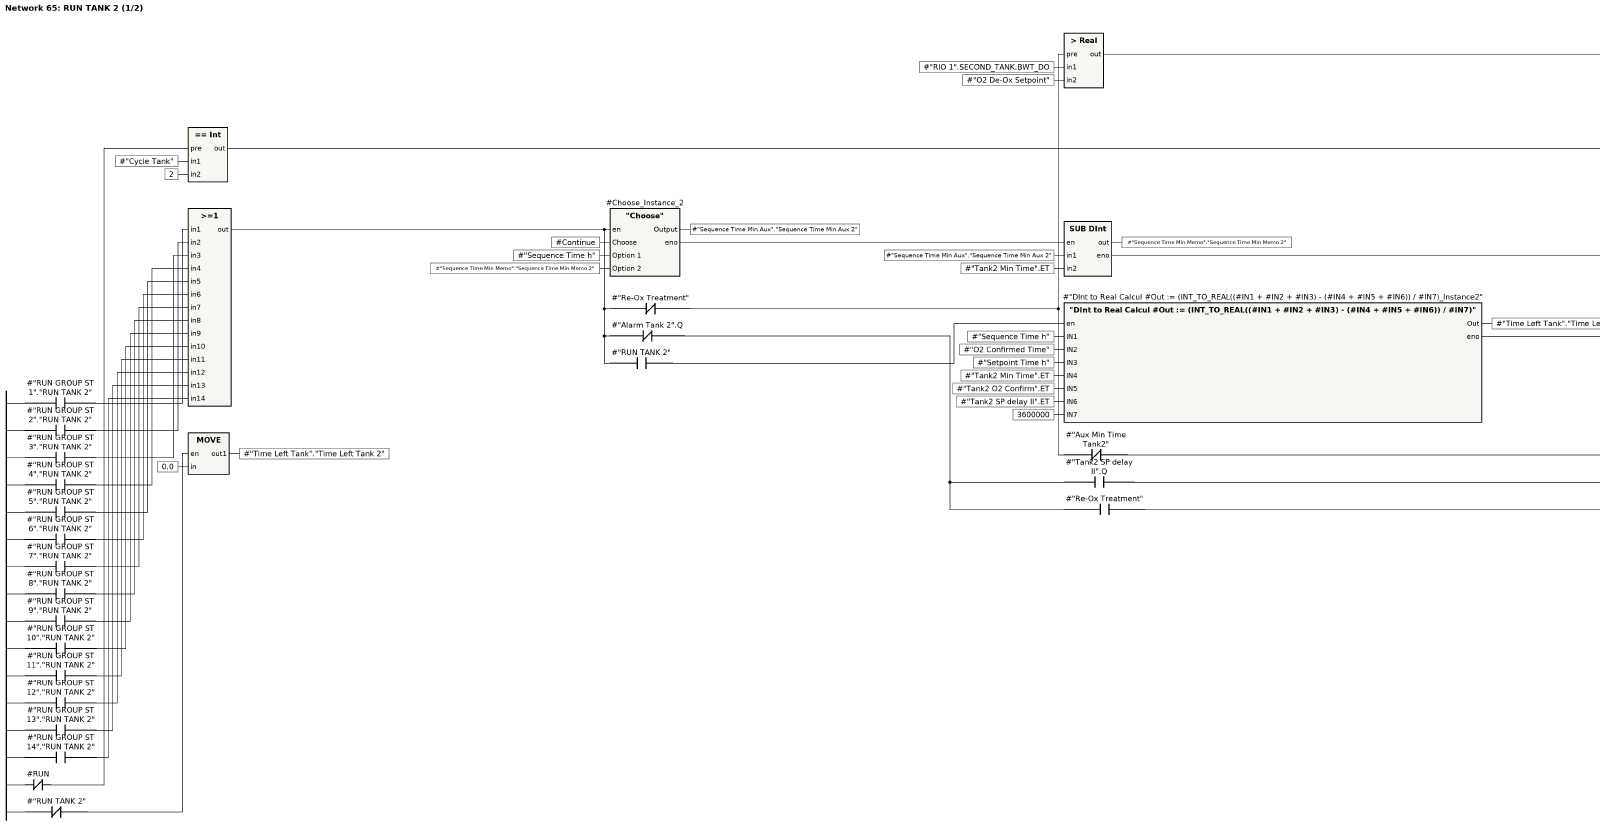
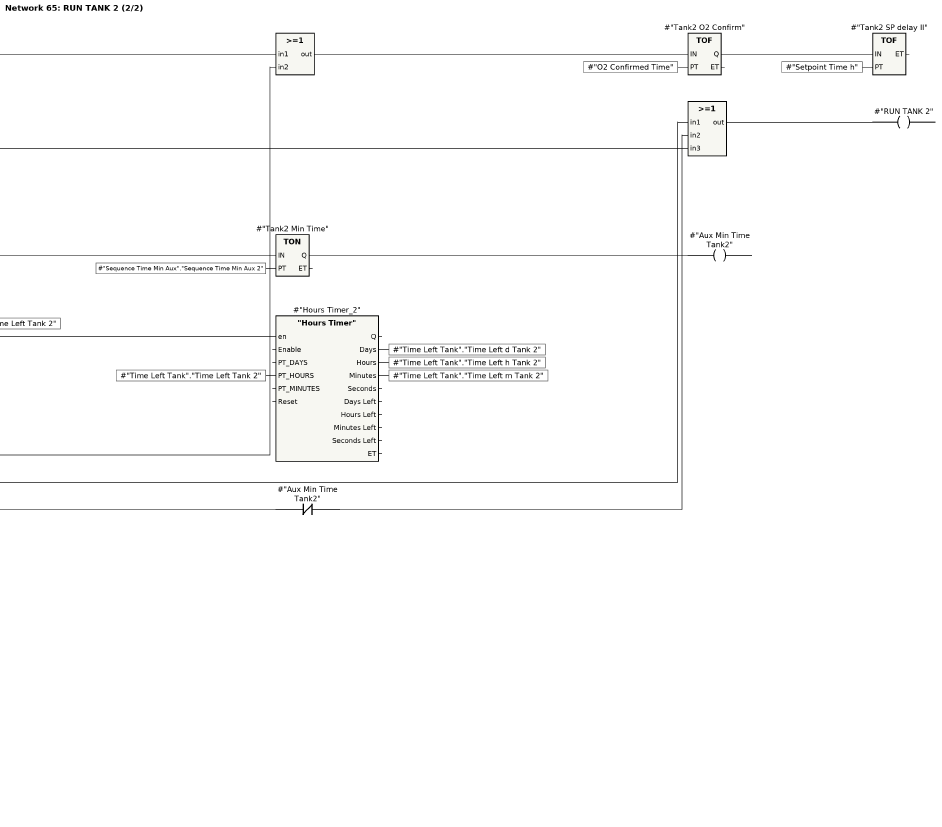
   #_w1 := #"RUN GROUP ST 1"."RUN TANK 2" OR #"RUN GROUP ST 2"."RUN TANK 2" OR #"RUN GROUP ST 3"."RUN TANK 2" OR #"RUN GROUP ST 4"."RUN TANK 2" OR #"RUN GROUP ST 5"."RUN TANK 2" OR #"RUN GROUP ST 6"."RUN TANK 2" OR #"RUN GROUP ST 7"."RUN TANK 2" OR #"RUN GROUP ST 8"."RUN TANK 2" OR #"RUN GROUP ST 9"."RUN TANK 2" OR #"RUN GROUP ST 10"."RUN TANK 2" OR #"RUN GROUP ST 11"."RUN TANK 2" OR #"RUN GROUP ST 12"."RUN TANK 2" OR #"RUN GROUP ST 13"."RUN TANK 2" OR #"RUN GROUP ST 14"."RUN TANK 2";
   #Choose_Instance_2(EN := #_w1,   // "Choose"
                      Choose := #Continue,
                      "Option 1" := #"Sequence Time h",
                      "Option 2" := #"Sequence Time Min Memo"."Sequence Time Min Memo 2",
                      Output => #"Sequence Time Min Aux"."Sequence Time Min Aux 2",
                      ENO => #_w2);
   IF #_w2 THEN
       #"Sequence Time Min Memo"."Sequence Time Min Memo 2" := #"Sequence Time Min Aux"."Sequence Time Min Aux 2" - #"Tank2 Min Time".ET;
   END_IF;
   #"Tank2 Min Time"(IN := #_w2, PT := #"Sequence Time Min Aux"."Sequence Time Min Aux 2");   // TON
   #"Aux Min Time Tank2" := #"Tank2 Min Time".Q;
   #"Tank2 O2 Confirm"(IN := #_w1 AND NOT #"Re-Ox Treatment" AND ((#"RIO 1".SECOND_TANK.BWT_DO > #"O2 De-Ox Setpoint") OR NOT #"Aux Min Time Tank2"),   // TOF
                       PT := #"O2 Confirmed Time");
   #"Tank2 SP delay II"(IN := #"Tank2 O2 Confirm".Q, PT := #"Setpoint Time h");   // TOF
   #"DInt to Real Calcul #Out := (INT_TO_REAL((#IN1 + #IN2 + #IN3) - (#IN4 + #IN5 + #IN6)) / #IN7)_Instance2"(EN := #_w1 AND #"RUN TANK 2",   // "DInt to Real Calcul #Out := (INT_TO_REAL((#IN1 + #IN2 + #IN3) - (#IN4 + #IN5 + #IN6)) / #IN7)"
                           IN1 := #"Sequence Time h",
                           IN2 := #"O2 Confirmed Time",
                           IN3 := #"Setpoint Time h",
                           IN4 := #"Tank2 Min Time".ET,
                           IN5 := #"Tank2 O2 Confirm".ET,
                           IN6 := #"Tank2 SP delay II".ET,
                           IN7 := 3600000,
                           Out => #"Time Left Tank"."Time Left Tank 2",
                           ENO => #_w3);
   IF #_w3 THEN
       #"Hours Timer_2"(PT_HOURS := #"Time Left Tank"."Time Left Tank 2",   // "Hours Timer"
                        Days => #"Time Left Tank"."Time Left d Tank 2",
                        Hours => #"Time Left Tank"."Time Left h Tank 2",
                        Minutes => #"Time Left Tank"."Time Left m Tank 2");
   END_IF;
   #"RUN TANK 2" := (#_w1 AND NOT #"Alarm Tank 2".Q AND (#"Tank2 SP delay II".Q OR (#"Re-Ox Treatment" AND NOT #"Aux Min Time Tank2"))) OR (NOT #RUN AND (#"Cycle Tank" = 2));
   IF NOT #"RUN TANK 2" THEN #"Time Left Tank"."Time Left Tank 2" := 0.0; END_IF;
END_REGION

REGION Network 66: RUN TANK 3
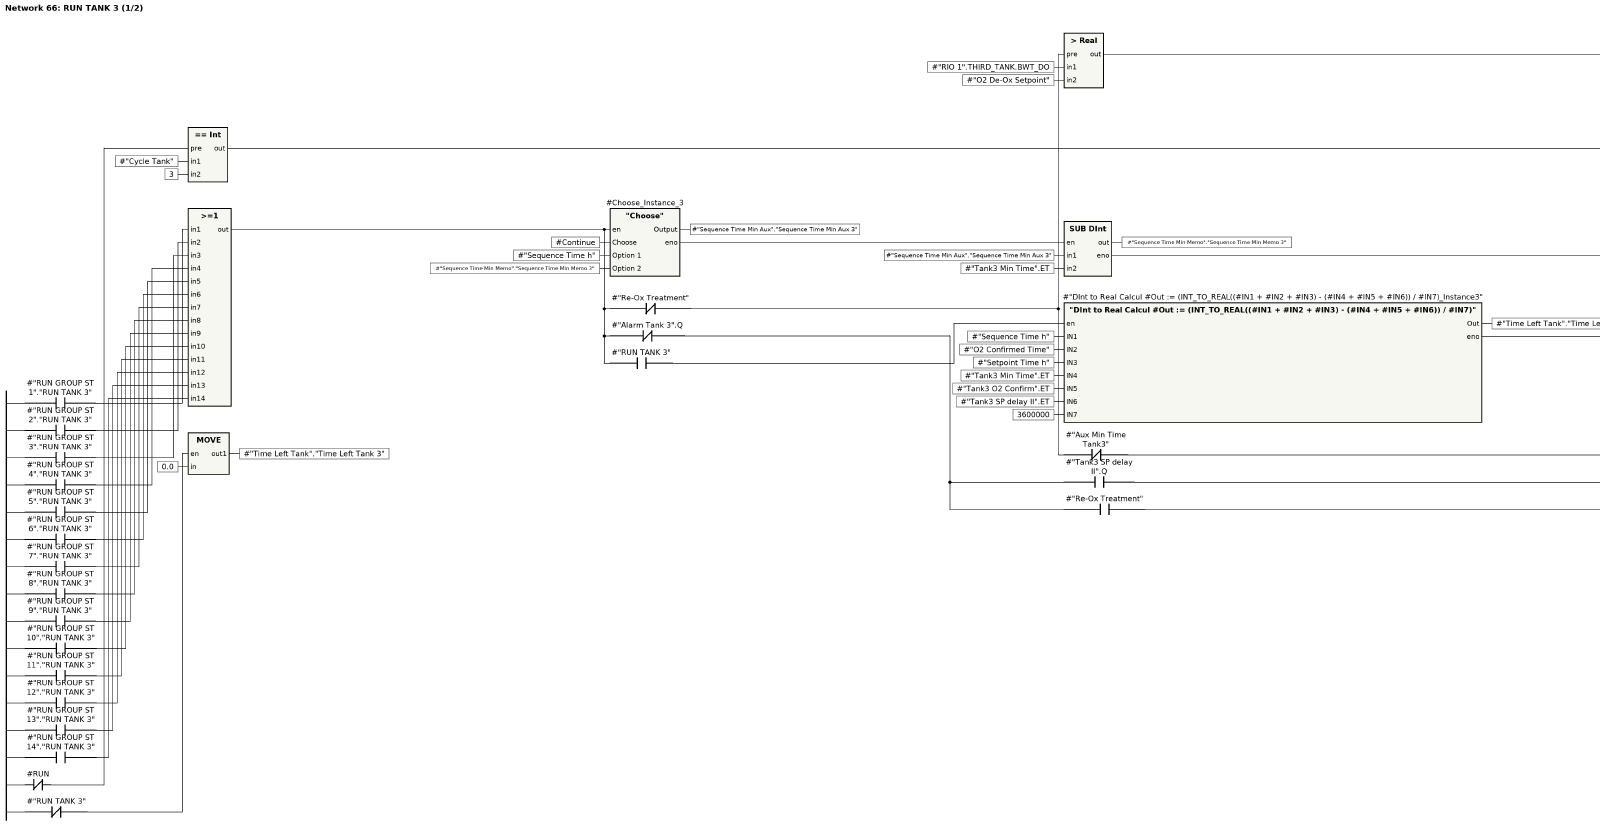
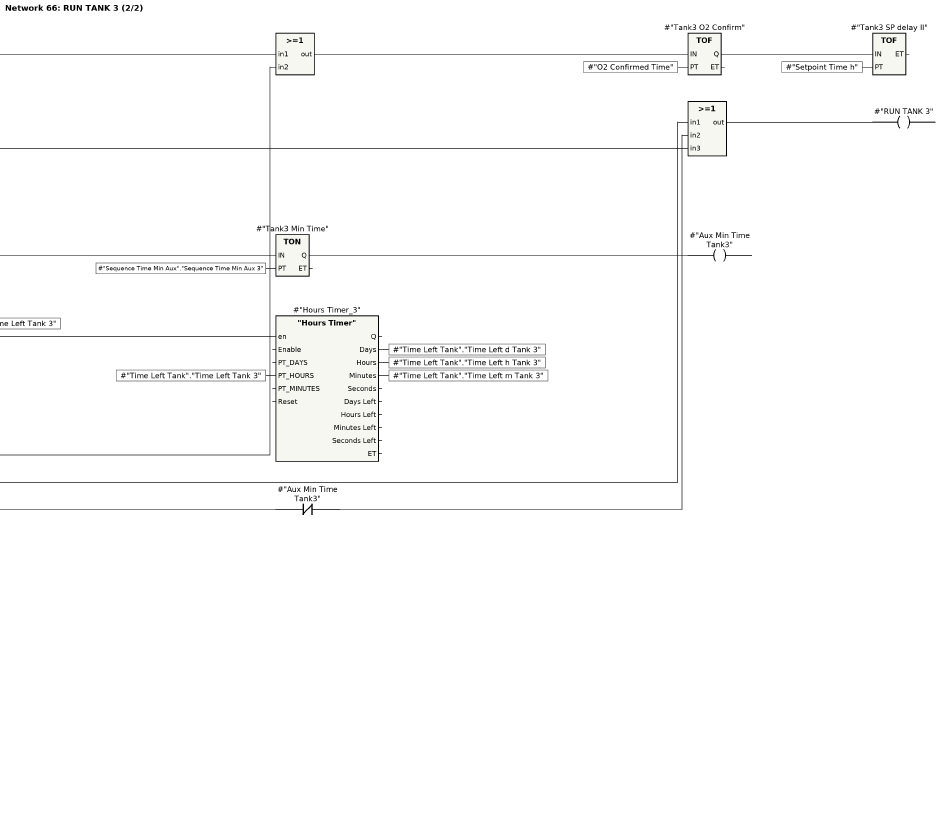
   #_w1 := #"RUN GROUP ST 1"."RUN TANK 3" OR #"RUN GROUP ST 2"."RUN TANK 3" OR #"RUN GROUP ST 3"."RUN TANK 3" OR #"RUN GROUP ST 4"."RUN TANK 3" OR #"RUN GROUP ST 5"."RUN TANK 3" OR #"RUN GROUP ST 6"."RUN TANK 3" OR #"RUN GROUP ST 7"."RUN TANK 3" OR #"RUN GROUP ST 8"."RUN TANK 3" OR #"RUN GROUP ST 9"."RUN TANK 3" OR #"RUN GROUP ST 10"."RUN TANK 3" OR #"RUN GROUP ST 11"."RUN TANK 3" OR #"RUN GROUP ST 12"."RUN TANK 3" OR #"RUN GROUP ST 13"."RUN TANK 3" OR #"RUN GROUP ST 14"."RUN TANK 3";
   #Choose_Instance_3(EN := #_w1,   // "Choose"
                      Choose := #Continue,
                      "Option 1" := #"Sequence Time h",
                      "Option 2" := #"Sequence Time Min Memo"."Sequence Time Min Memo 3",
                      Output => #"Sequence Time Min Aux"."Sequence Time Min Aux 3",
                      ENO => #_w2);
   IF #_w2 THEN
       #"Sequence Time Min Memo"."Sequence Time Min Memo 3" := #"Sequence Time Min Aux"."Sequence Time Min Aux 3" - #"Tank3 Min Time".ET;   // Memory of remained time for use to continue
   END_IF;
   #"Tank3 Min Time"(IN := #_w2, PT := #"Sequence Time Min Aux"."Sequence Time Min Aux 3");   // TON
   #"Aux Min Time Tank3" := #"Tank3 Min Time".Q;
   #"Tank3 O2 Confirm"(IN := #_w1 AND NOT #"Re-Ox Treatment" AND ((#"RIO 1".THIRD_TANK.BWT_DO > #"O2 De-Ox Setpoint") OR NOT #"Aux Min Time Tank3"),   // TOF
                       PT := #"O2 Confirmed Time");
   #"Tank3 SP delay II"(IN := #"Tank3 O2 Confirm".Q, PT := #"Setpoint Time h");   // TOF
   #"DInt to Real Calcul #Out := (INT_TO_REAL((#IN1 + #IN2 + #IN3) - (#IN4 + #IN5 + #IN6)) / #IN7)_Instance3"(EN := #_w1 AND #"RUN TANK 3",   // "DInt to Real Calcul #Out := (INT_TO_REAL((#IN1 + #IN2 + #IN3) - (#IN4 + #IN5 + #IN6)) / #IN7)"
                           IN1 := #"Sequence Time h",
                           IN2 := #"O2 Confirmed Time",
                           IN3 := #"Setpoint Time h",
                           IN4 := #"Tank3 Min Time".ET,
                           IN5 := #"Tank3 O2 Confirm".ET,
                           IN6 := #"Tank3 SP delay II".ET,
                           IN7 := 3600000,
                           Out => #"Time Left Tank"."Time Left Tank 3",
                           ENO => #_w3);
   IF #_w3 THEN
       #"Hours Timer_3"(PT_HOURS := #"Time Left Tank"."Time Left Tank 3",   // "Hours Timer"
                        Days => #"Time Left Tank"."Time Left d Tank 3",
                        Hours => #"Time Left Tank"."Time Left h Tank 3",
                        Minutes => #"Time Left Tank"."Time Left m Tank 3");
   END_IF;
   #"RUN TANK 3" := (#_w1 AND NOT #"Alarm Tank 3".Q AND (#"Tank3 SP delay II".Q OR (#"Re-Ox Treatment" AND NOT #"Aux Min Time Tank3"))) OR (NOT #RUN AND (#"Cycle Tank" = 3));
   IF NOT #"RUN TANK 3" THEN #"Time Left Tank"."Time Left Tank 3" := 0.0; END_IF;
END_REGION

REGION Network 67: RUN TANK 4
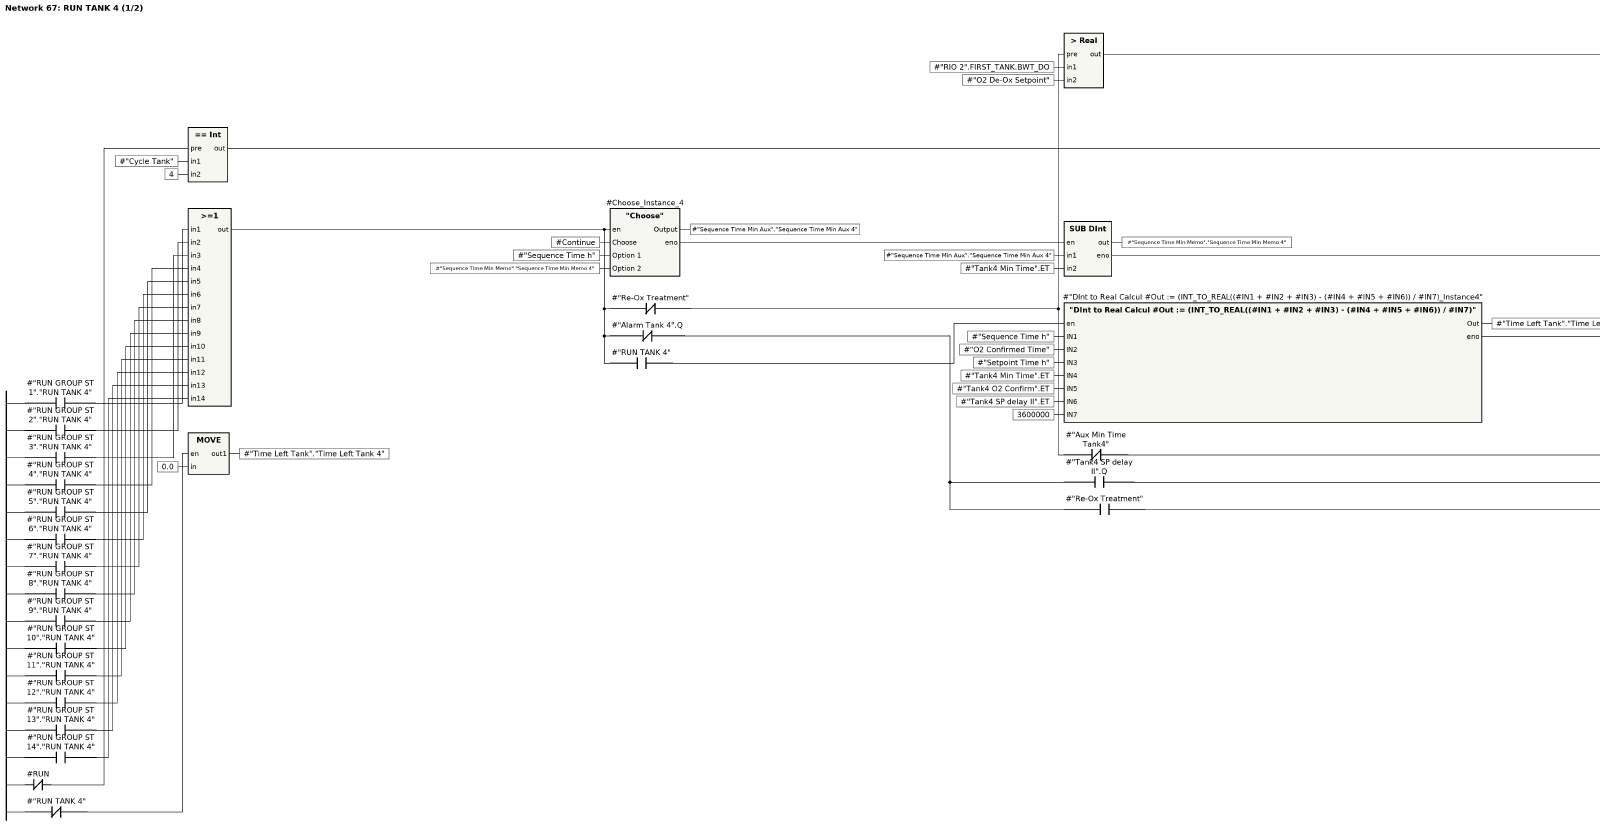
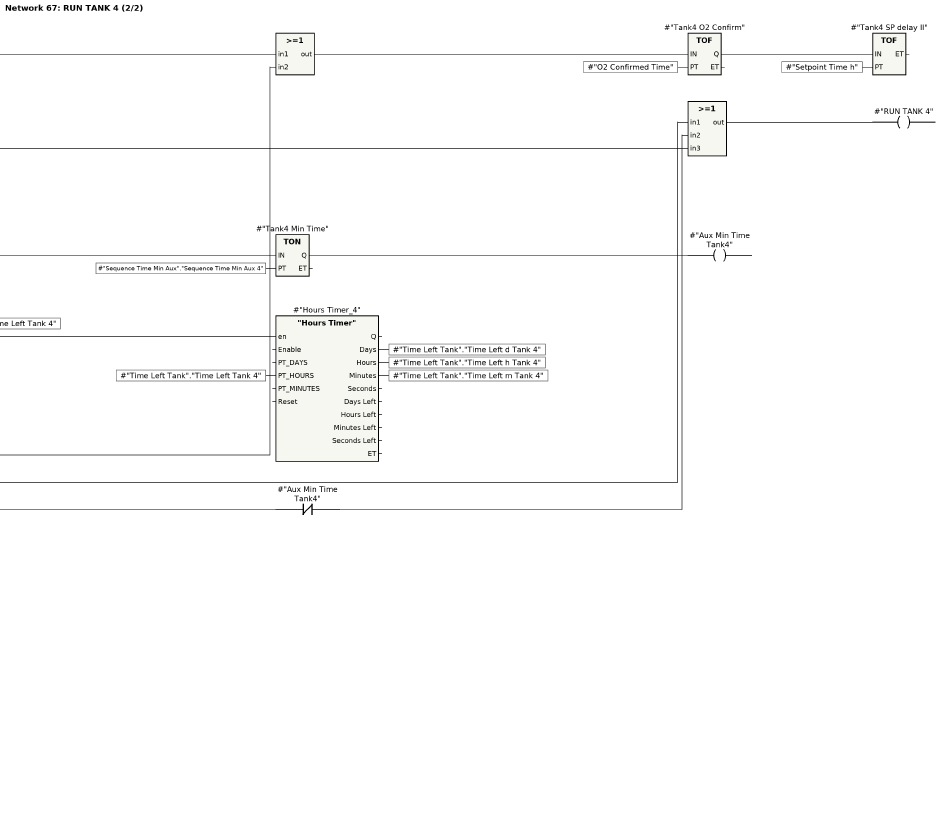
   #_w1 := #"RUN GROUP ST 1"."RUN TANK 4" OR #"RUN GROUP ST 2"."RUN TANK 4" OR #"RUN GROUP ST 3"."RUN TANK 4" OR #"RUN GROUP ST 4"."RUN TANK 4" OR #"RUN GROUP ST 5"."RUN TANK 4" OR #"RUN GROUP ST 6"."RUN TANK 4" OR #"RUN GROUP ST 7"."RUN TANK 4" OR #"RUN GROUP ST 8"."RUN TANK 4" OR #"RUN GROUP ST 9"."RUN TANK 4" OR #"RUN GROUP ST 10"."RUN TANK 4" OR #"RUN GROUP ST 11"."RUN TANK 4" OR #"RUN GROUP ST 12"."RUN TANK 4" OR #"RUN GROUP ST 13"."RUN TANK 4" OR #"RUN GROUP ST 14"."RUN TANK 4";
   #Choose_Instance_4(EN := #_w1,   // "Choose"
                      Choose := #Continue,
                      "Option 1" := #"Sequence Time h",
                      "Option 2" := #"Sequence Time Min Memo"."Sequence Time Min Memo 4",
                      Output => #"Sequence Time Min Aux"."Sequence Time Min Aux 4",
                      ENO => #_w2);
   IF #_w2 THEN
       #"Sequence Time Min Memo"."Sequence Time Min Memo 4" := #"Sequence Time Min Aux"."Sequence Time Min Aux 4" - #"Tank4 Min Time".ET;   // Memory of remained time for use to continue
   END_IF;
   #"Tank4 Min Time"(IN := #_w2, PT := #"Sequence Time Min Aux"."Sequence Time Min Aux 4");   // TON
   #"Aux Min Time Tank4" := #"Tank4 Min Time".Q;
   #"Tank4 O2 Confirm"(IN := #_w1 AND NOT #"Re-Ox Treatment" AND ((#"RIO 2".FIRST_TANK.BWT_DO > #"O2 De-Ox Setpoint") OR NOT #"Aux Min Time Tank4"),   // TOF
                       PT := #"O2 Confirmed Time");
   #"Tank4 SP delay II"(IN := #"Tank4 O2 Confirm".Q, PT := #"Setpoint Time h");   // TOF
   #"DInt to Real Calcul #Out := (INT_TO_REAL((#IN1 + #IN2 + #IN3) - (#IN4 + #IN5 + #IN6)) / #IN7)_Instance4"(EN := #_w1 AND #"RUN TANK 4",   // "DInt to Real Calcul #Out := (INT_TO_REAL((#IN1 + #IN2 + #IN3) - (#IN4 + #IN5 + #IN6)) / #IN7)"
                           IN1 := #"Sequence Time h",
                           IN2 := #"O2 Confirmed Time",
                           IN3 := #"Setpoint Time h",
                           IN4 := #"Tank4 Min Time".ET,
                           IN5 := #"Tank4 O2 Confirm".ET,
                           IN6 := #"Tank4 SP delay II".ET,
                           IN7 := 3600000,
                           Out => #"Time Left Tank"."Time Left Tank 4",
                           ENO => #_w3);
   IF #_w3 THEN
       #"Hours Timer_4"(PT_HOURS := #"Time Left Tank"."Time Left Tank 4",   // "Hours Timer"
                        Days => #"Time Left Tank"."Time Left d Tank 4",
                        Hours => #"Time Left Tank"."Time Left h Tank 4",
                        Minutes => #"Time Left Tank"."Time Left m Tank 4");
   END_IF;
   #"RUN TANK 4" := (#_w1 AND NOT #"Alarm Tank 4".Q AND (#"Tank4 SP delay II".Q OR (#"Re-Ox Treatment" AND NOT #"Aux Min Time Tank4"))) OR (NOT #RUN AND (#"Cycle Tank" = 4));
   IF NOT #"RUN TANK 4" THEN #"Time Left Tank"."Time Left Tank 4" := 0.0; END_IF;
END_REGION

REGION Network 68: RUN TANK 5
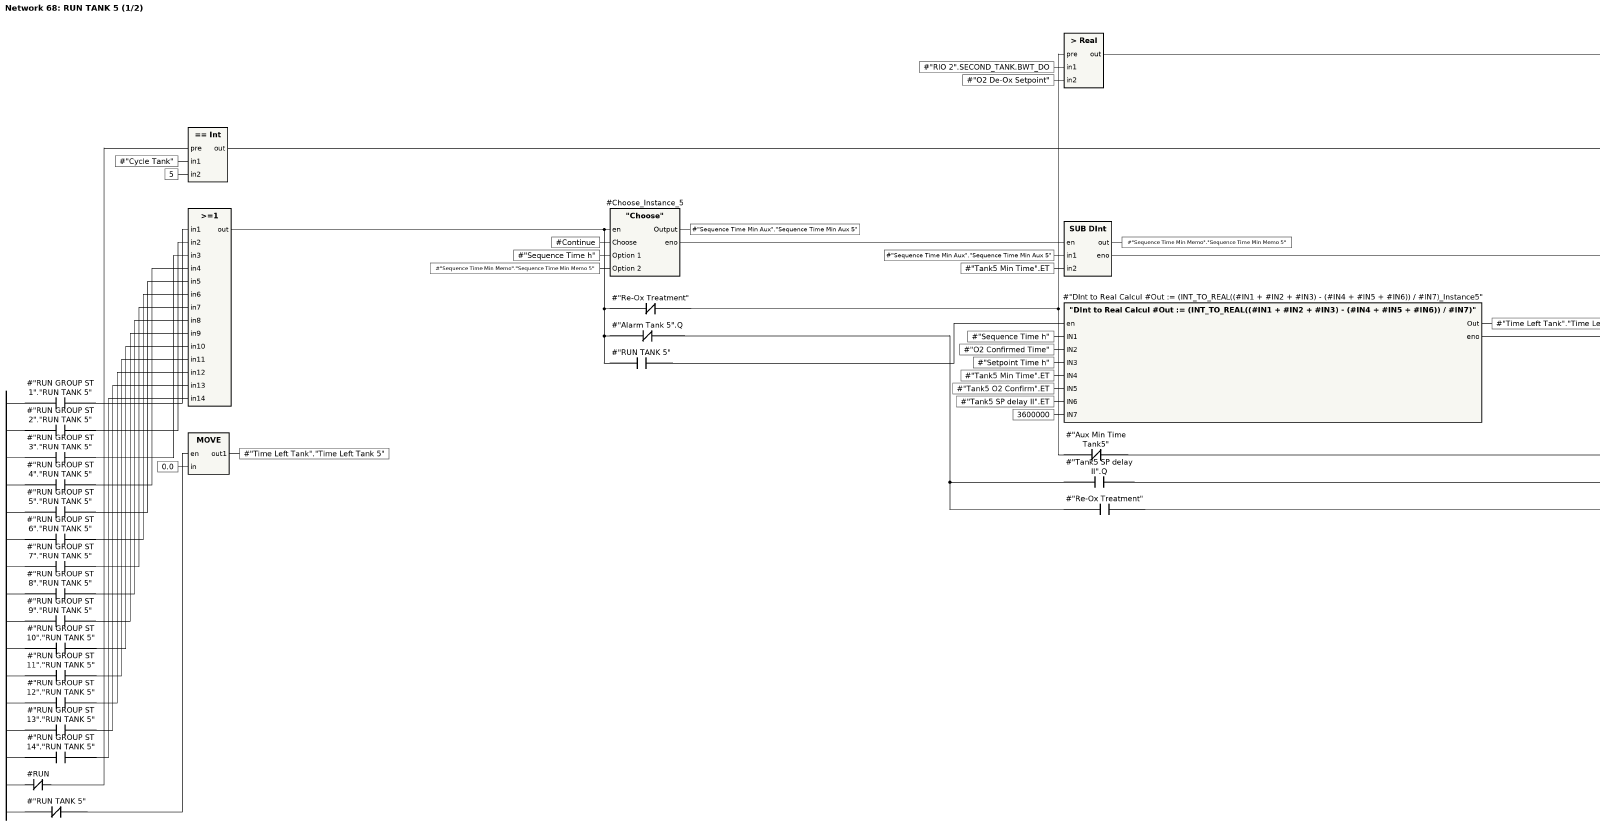
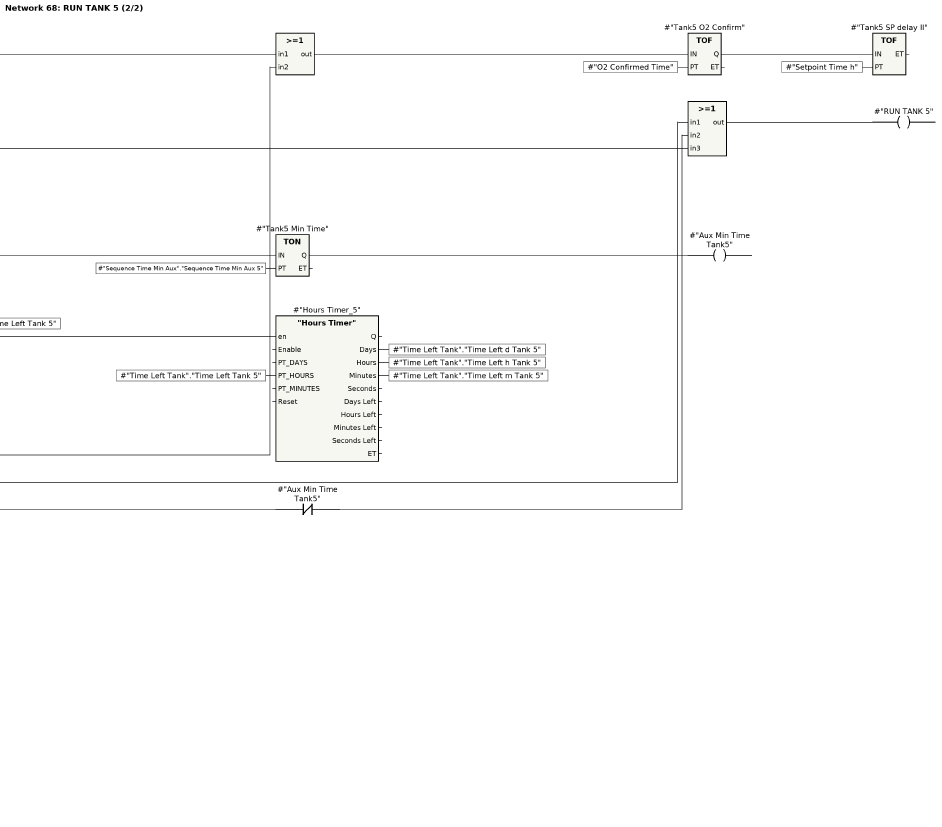
   #_w1 := #"RUN GROUP ST 1"."RUN TANK 5" OR #"RUN GROUP ST 2"."RUN TANK 5" OR #"RUN GROUP ST 3"."RUN TANK 5" OR #"RUN GROUP ST 4"."RUN TANK 5" OR #"RUN GROUP ST 5"."RUN TANK 5" OR #"RUN GROUP ST 6"."RUN TANK 5" OR #"RUN GROUP ST 7"."RUN TANK 5" OR #"RUN GROUP ST 8"."RUN TANK 5" OR #"RUN GROUP ST 9"."RUN TANK 5" OR #"RUN GROUP ST 10"."RUN TANK 5" OR #"RUN GROUP ST 11"."RUN TANK 5" OR #"RUN GROUP ST 12"."RUN TANK 5" OR #"RUN GROUP ST 13"."RUN TANK 5" OR #"RUN GROUP ST 14"."RUN TANK 5";
   #Choose_Instance_5(EN := #_w1,   // "Choose"
                      Choose := #Continue,
                      "Option 1" := #"Sequence Time h",
                      "Option 2" := #"Sequence Time Min Memo"."Sequence Time Min Memo 5",
                      Output => #"Sequence Time Min Aux"."Sequence Time Min Aux 5",
                      ENO => #_w2);
   IF #_w2 THEN
       #"Sequence Time Min Memo"."Sequence Time Min Memo 5" := #"Sequence Time Min Aux"."Sequence Time Min Aux 5" - #"Tank5 Min Time".ET;   // Memory of remained time for use to continue
   END_IF;
   #"Tank5 Min Time"(IN := #_w2, PT := #"Sequence Time Min Aux"."Sequence Time Min Aux 5");   // TON
   #"Aux Min Time Tank5" := #"Tank5 Min Time".Q;
   #"Tank5 O2 Confirm"(IN := #_w1 AND NOT #"Re-Ox Treatment" AND ((#"RIO 2".SECOND_TANK.BWT_DO > #"O2 De-Ox Setpoint") OR NOT #"Aux Min Time Tank5"),   // TOF
                       PT := #"O2 Confirmed Time");
   #"Tank5 SP delay II"(IN := #"Tank5 O2 Confirm".Q, PT := #"Setpoint Time h");   // TOF
   #"DInt to Real Calcul #Out := (INT_TO_REAL((#IN1 + #IN2 + #IN3) - (#IN4 + #IN5 + #IN6)) / #IN7)_Instance5"(EN := #_w1 AND #"RUN TANK 5",   // "DInt to Real Calcul #Out := (INT_TO_REAL((#IN1 + #IN2 + #IN3) - (#IN4 + #IN5 + #IN6)) / #IN7)"
                           IN1 := #"Sequence Time h",
                           IN2 := #"O2 Confirmed Time",
                           IN3 := #"Setpoint Time h",
                           IN4 := #"Tank5 Min Time".ET,
                           IN5 := #"Tank5 O2 Confirm".ET,
                           IN6 := #"Tank5 SP delay II".ET,
                           IN7 := 3600000,
                           Out => #"Time Left Tank"."Time Left Tank 5",
                           ENO => #_w3);
   IF #_w3 THEN
       #"Hours Timer_5"(PT_HOURS := #"Time Left Tank"."Time Left Tank 5",   // "Hours Timer"
                        Days => #"Time Left Tank"."Time Left d Tank 5",
                        Hours => #"Time Left Tank"."Time Left h Tank 5",
                        Minutes => #"Time Left Tank"."Time Left m Tank 5");
   END_IF;
   #"RUN TANK 5" := (#_w1 AND NOT #"Alarm Tank 5".Q AND (#"Tank5 SP delay II".Q OR (#"Re-Ox Treatment" AND NOT #"Aux Min Time Tank5"))) OR (NOT #RUN AND (#"Cycle Tank" = 5));
   IF NOT #"RUN TANK 5" THEN #"Time Left Tank"."Time Left Tank 5" := 0.0; END_IF;
END_REGION

REGION Network 69: RUN TANK 6
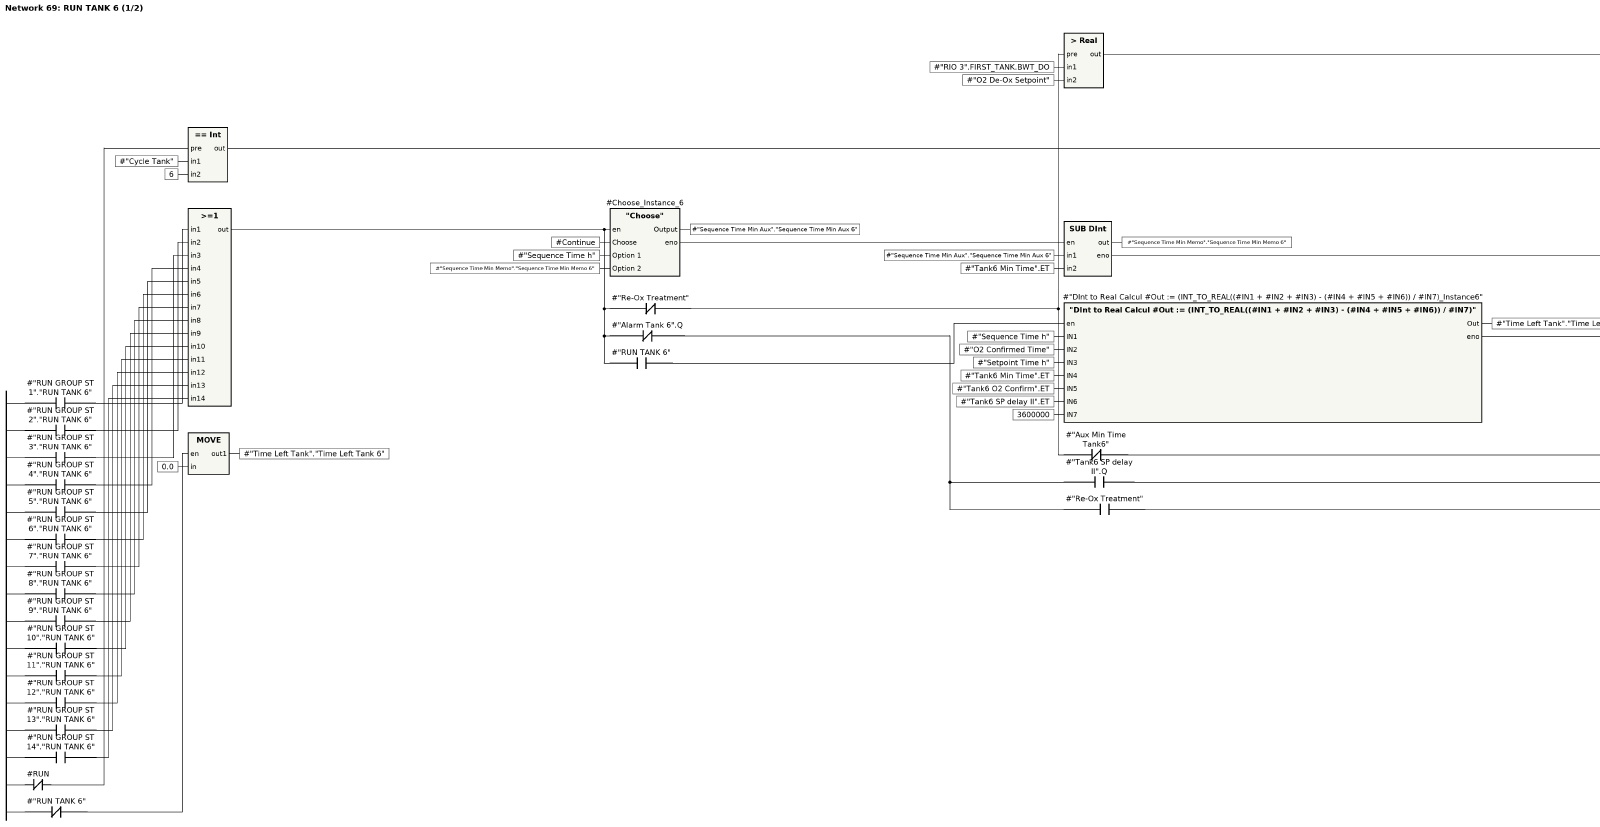
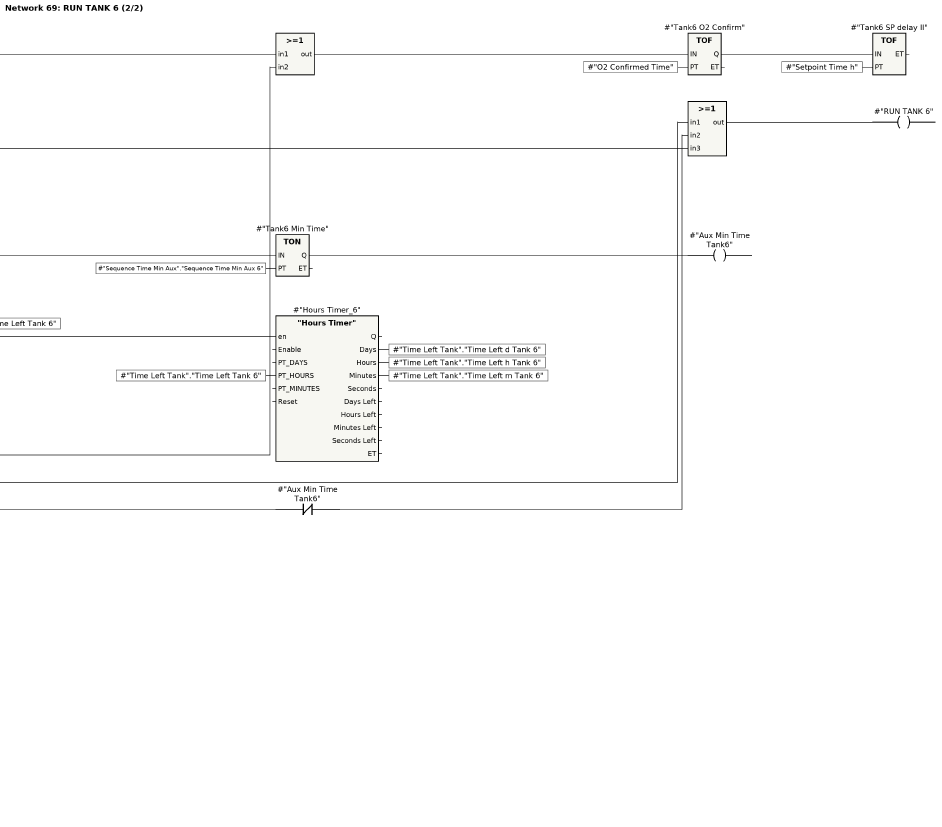
   #_w1 := #"RUN GROUP ST 1"."RUN TANK 6" OR #"RUN GROUP ST 2"."RUN TANK 6" OR #"RUN GROUP ST 3"."RUN TANK 6" OR #"RUN GROUP ST 4"."RUN TANK 6" OR #"RUN GROUP ST 5"."RUN TANK 6" OR #"RUN GROUP ST 6"."RUN TANK 6" OR #"RUN GROUP ST 7"."RUN TANK 6" OR #"RUN GROUP ST 8"."RUN TANK 6" OR #"RUN GROUP ST 9"."RUN TANK 6" OR #"RUN GROUP ST 10"."RUN TANK 6" OR #"RUN GROUP ST 11"."RUN TANK 6" OR #"RUN GROUP ST 12"."RUN TANK 6" OR #"RUN GROUP ST 13"."RUN TANK 6" OR #"RUN GROUP ST 14"."RUN TANK 6";
   #Choose_Instance_6(EN := #_w1,   // "Choose"
                      Choose := #Continue,
                      "Option 1" := #"Sequence Time h",
                      "Option 2" := #"Sequence Time Min Memo"."Sequence Time Min Memo 6",
                      Output => #"Sequence Time Min Aux"."Sequence Time Min Aux 6",
                      ENO => #_w2);
   IF #_w2 THEN
       #"Sequence Time Min Memo"."Sequence Time Min Memo 6" := #"Sequence Time Min Aux"."Sequence Time Min Aux 6" - #"Tank6 Min Time".ET;   // Memory of remained time for use to continue
   END_IF;
   #"Tank6 Min Time"(IN := #_w2, PT := #"Sequence Time Min Aux"."Sequence Time Min Aux 6");   // TON
   #"Aux Min Time Tank6" := #"Tank6 Min Time".Q;
   #"Tank6 O2 Confirm"(IN := #_w1 AND NOT #"Re-Ox Treatment" AND ((#"RIO 3".FIRST_TANK.BWT_DO > #"O2 De-Ox Setpoint") OR NOT #"Aux Min Time Tank6"),   // TOF
                       PT := #"O2 Confirmed Time");
   #"Tank6 SP delay II"(IN := #"Tank6 O2 Confirm".Q, PT := #"Setpoint Time h");   // TOF
   #"DInt to Real Calcul #Out := (INT_TO_REAL((#IN1 + #IN2 + #IN3) - (#IN4 + #IN5 + #IN6)) / #IN7)_Instance6"(EN := #_w1 AND #"RUN TANK 6",   // "DInt to Real Calcul #Out := (INT_TO_REAL((#IN1 + #IN2 + #IN3) - (#IN4 + #IN5 + #IN6)) / #IN7)"
                           IN1 := #"Sequence Time h",
                           IN2 := #"O2 Confirmed Time",
                           IN3 := #"Setpoint Time h",
                           IN4 := #"Tank6 Min Time".ET,
                           IN5 := #"Tank6 O2 Confirm".ET,
                           IN6 := #"Tank6 SP delay II".ET,
                           IN7 := 3600000,
                           Out => #"Time Left Tank"."Time Left Tank 6",
                           ENO => #_w3);
   IF #_w3 THEN
       #"Hours Timer_6"(PT_HOURS := #"Time Left Tank"."Time Left Tank 6",   // "Hours Timer"
                        Days => #"Time Left Tank"."Time Left d Tank 6",
                        Hours => #"Time Left Tank"."Time Left h Tank 6",
                        Minutes => #"Time Left Tank"."Time Left m Tank 6");
   END_IF;
   #"RUN TANK 6" := (#_w1 AND NOT #"Alarm Tank 6".Q AND (#"Tank6 SP delay II".Q OR (#"Re-Ox Treatment" AND NOT #"Aux Min Time Tank6"))) OR (NOT #RUN AND (#"Cycle Tank" = 6));
   IF NOT #"RUN TANK 6" THEN #"Time Left Tank"."Time Left Tank 6" := 0.0; END_IF;
END_REGION

REGION Network 70: RUN TANK 7
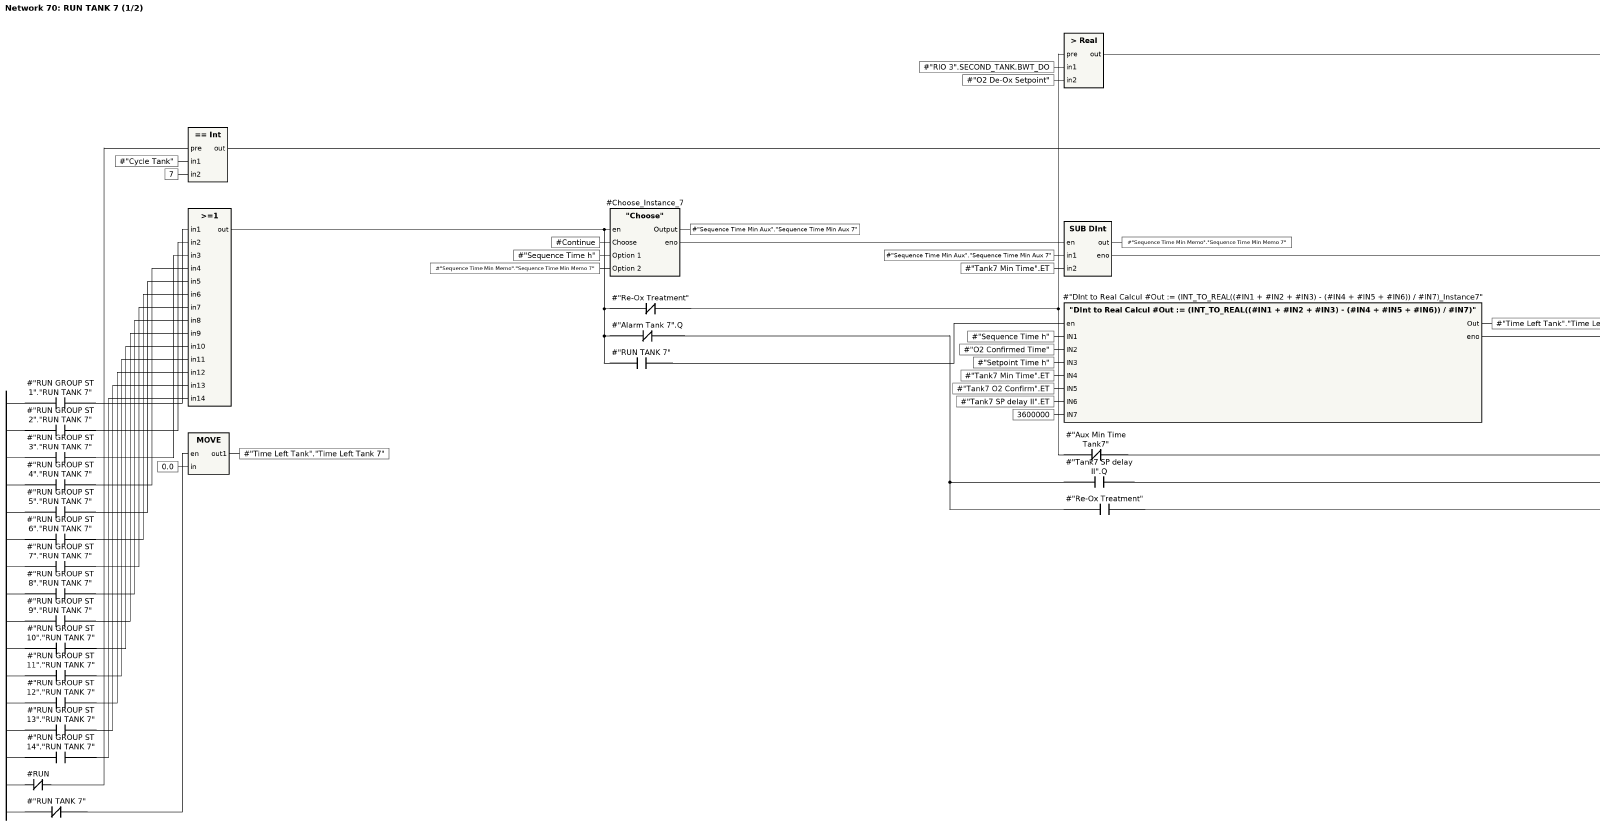
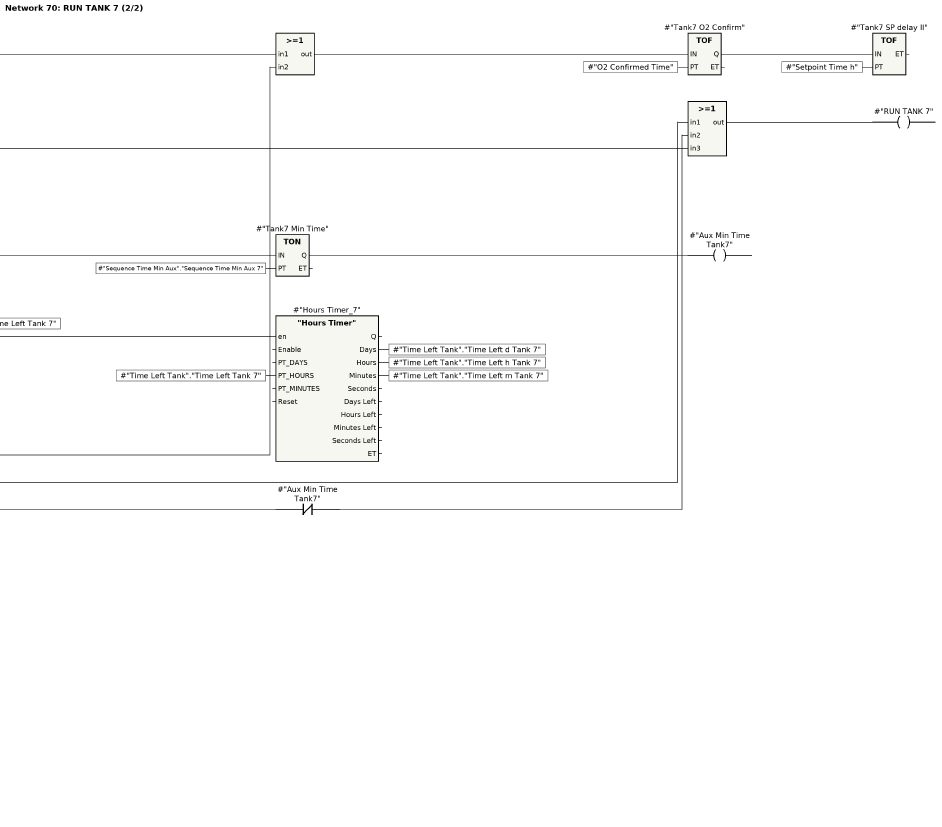
   #_w1 := #"RUN GROUP ST 1"."RUN TANK 7" OR #"RUN GROUP ST 2"."RUN TANK 7" OR #"RUN GROUP ST 3"."RUN TANK 7" OR #"RUN GROUP ST 4"."RUN TANK 7" OR #"RUN GROUP ST 5"."RUN TANK 7" OR #"RUN GROUP ST 6"."RUN TANK 7" OR #"RUN GROUP ST 7"."RUN TANK 7" OR #"RUN GROUP ST 8"."RUN TANK 7" OR #"RUN GROUP ST 9"."RUN TANK 7" OR #"RUN GROUP ST 10"."RUN TANK 7" OR #"RUN GROUP ST 11"."RUN TANK 7" OR #"RUN GROUP ST 12"."RUN TANK 7" OR #"RUN GROUP ST 13"."RUN TANK 7" OR #"RUN GROUP ST 14"."RUN TANK 7";
   #Choose_Instance_7(EN := #_w1,   // "Choose"
                      Choose := #Continue,
                      "Option 1" := #"Sequence Time h",
                      "Option 2" := #"Sequence Time Min Memo"."Sequence Time Min Memo 7",
                      Output => #"Sequence Time Min Aux"."Sequence Time Min Aux 7",
                      ENO => #_w2);
   IF #_w2 THEN
       #"Sequence Time Min Memo"."Sequence Time Min Memo 7" := #"Sequence Time Min Aux"."Sequence Time Min Aux 7" - #"Tank7 Min Time".ET;   // Memory of remained time for use to continue
   END_IF;
   #"Tank7 Min Time"(IN := #_w2, PT := #"Sequence Time Min Aux"."Sequence Time Min Aux 7");   // TON
   #"Aux Min Time Tank7" := #"Tank7 Min Time".Q;
   #"Tank7 O2 Confirm"(IN := #_w1 AND NOT #"Re-Ox Treatment" AND ((#"RIO 3".SECOND_TANK.BWT_DO > #"O2 De-Ox Setpoint") OR NOT #"Aux Min Time Tank7"),   // TOF
                       PT := #"O2 Confirmed Time");
   #"Tank7 SP delay II"(IN := #"Tank7 O2 Confirm".Q, PT := #"Setpoint Time h");   // TOF
   #"DInt to Real Calcul #Out := (INT_TO_REAL((#IN1 + #IN2 + #IN3) - (#IN4 + #IN5 + #IN6)) / #IN7)_Instance7"(EN := #_w1 AND #"RUN TANK 7",   // "DInt to Real Calcul #Out := (INT_TO_REAL((#IN1 + #IN2 + #IN3) - (#IN4 + #IN5 + #IN6)) / #IN7)"
                           IN1 := #"Sequence Time h",
                           IN2 := #"O2 Confirmed Time",
                           IN3 := #"Setpoint Time h",
                           IN4 := #"Tank7 Min Time".ET,
                           IN5 := #"Tank7 O2 Confirm".ET,
                           IN6 := #"Tank7 SP delay II".ET,
                           IN7 := 3600000,
                           Out => #"Time Left Tank"."Time Left Tank 7",
                           ENO => #_w3);
   IF #_w3 THEN
       #"Hours Timer_7"(PT_HOURS := #"Time Left Tank"."Time Left Tank 7",   // "Hours Timer"
                        Days => #"Time Left Tank"."Time Left d Tank 7",
                        Hours => #"Time Left Tank"."Time Left h Tank 7",
                        Minutes => #"Time Left Tank"."Time Left m Tank 7");
   END_IF;
   #"RUN TANK 7" := (#_w1 AND NOT #"Alarm Tank 7".Q AND (#"Tank7 SP delay II".Q OR (#"Re-Ox Treatment" AND NOT #"Aux Min Time Tank7"))) OR (NOT #RUN AND (#"Cycle Tank" = 7));
   IF NOT #"RUN TANK 7" THEN #"Time Left Tank"."Time Left Tank 7" := 0.0; END_IF;
END_REGION

REGION Network 71: RUN TANK 8